REGION Network 2: Dose_Control_Linie_1
   IF "GDB_PLC".Start_Modus_Linie_1 AND NOT "GDB_PLC".Stop_Modus_Linie_1 THEN
       "FB_Dose_Control_DB_1"(Trigger_Start := "GDB_PLC".Dosierung_Start_Linie_1,   // "FB_Dose_Control"
                              Flow_Raw := "Tank 2 (Flow Meter)",
                              Target_Volume := "GDB_Getränk".Getränk_Linie_1.Dosiervolumen,
                              Not_Aus := "GDB_PLC".Not_Aus_Modus,
                              Discharge_Valve => "Tank 2 (Discharge Valve)",
                              Dosing_Status => "GDB_PLC".Dosing_Activate_Linie_1,
                              Füllmenge => "GDB_HMI".Füllmenge_Linie_1);
   END_IF;
END_REGION
END_ORGANIZATION_BLOCK

(* ===== HMI "HMI_RT_1" =====
system functions are stored by id; their names below are inferred from use
connection "HMI_Verbindung_1": ETHERNET, SMART_S7_1200_OMS

HMI tags "Standard-Variablentabelle"
   "Variable_Bildnummer" : UInt, internal
   "Start Button 1" : Bool = PLC "Start Button 1" AT %I5.0, 100 ms
   "Start Button 1 (Light)" : Bool = PLC "Start Button 1 (Light)" AT %Q4.4, 100 ms
   "Stop Button 1" : Bool = PLC "Stop Button 1" AT %I5.2, 100 ms
   "Emergency Stop 1" : Bool = PLC "Emergency Stop 1" AT %I3.7, 100 ms
   "GDB_PLC_Start_Modus" : Bool = PLC GDB_PLC.Start_Modus_Hauptleitung, 100 ms
   "GDB_PLC_Not_Aus_Modus" : Bool = PLC GDB_PLC.Not_Aus_Modus, 100 ms
   "GDB_HMI_Füllmenge" : Real = PLC GDB_HMI.Füllmenge_Linie_0, 100 ms
   "GDB_PLC_Dosing_Activate" : Bool = PLC GDB_PLC.Dosing_Activate_Linie_0, 100 ms
   "GDB_PLC_Füllventil_Stand" : Bool = PLC GDB_PLC.Füllventil_closed_Linie_0, 100 ms
   "Stop Button 1 (Light)" : Bool = PLC "Stop Button 1 (Light)" AT %Q4.6, 100 ms
   "GDB_HMI_Reset_Gesamtteile_0" : Bool = PLC GDB_HMI.Reset_Gesamtteile_0, 100 ms
   "GDB_HMI_Reset_Ausschluss_0" : Bool = PLC GDB_HMI.Reset_Ausschluss_0, 100 ms
   "GDB_PLC_Gesamtteile_Linie_0" : Int = PLC GDB_PLC.Gesamtteile_Linie_0, 100 ms
   "GDB_PLC_Altuell_Gewicht_Linie_0" : Real = PLC GDB_PLC.Altuell_Gewicht_Linie_0, 100 ms
   "GDB_PLC_Tankfüllvolumen" : Real = PLC GDB_PLC.Tankfüllvolumen_0, 100 ms
   "GDB_PLC_Dosiervolumen" : Real = PLC GDB_PLC.Dosiervolumen_0, 100 ms
   "GDB_Getränk_Getränk_Linie_1_VAR_Rezeptur_Datensatz" : Int = PLC GDB_Getränk.Getränk_Linie_1.VAR_Rezeptur_Datensatz, 100 ms
   "GDB_Getränk_Getränk_Linie_0_VAR_Rezeptur_Datensatz" : Int = PLC GDB_Getränk.Getränk_Linie_0.VAR_Rezeptur_Datensatz, 100 ms
   "GDB_Getränk_Getränk_Linie_0_VAR_Rezeptur" : Int = PLC GDB_Getränk.Getränk_Linie_0.VAR_Rezeptur, 100 ms
   "GDB_Getränk_Getränk_Linie_0_Tankfüllvolumen" : Real = PLC GDB_Getränk.Getränk_Linie_0.Tankfüllvolumen, 100 ms
   "GDB_Getränk_Getränk_Linie_0_Dosiervolumen" : Real = PLC GDB_Getränk.Getränk_Linie_0.Dosiervolumen, 100 ms
   "GDB_PLC_Tank_1_Level_norm" : Real = PLC GDB_PLC.Tank_1_Level_norm, 100 ms
   "Start Button 0" : Bool = PLC "Start Button 0" AT %I5.3, 100 ms
   "Stop Button 0" : Bool = PLC "Stop Button 0" AT %I5.1, 100 ms
   "Emergency Stop 0" : Bool = PLC "Emergency Stop 0" AT %I3.6, 100 ms
   "GDB_Getränk_Getränk_Linie_1_Tankfüllvolumen" : Real = PLC GDB_Getränk.Getränk_Linie_1.Tankfüllvolumen, 100 ms
   "GDB_Getränk_Getränk_Linie_1_Dosiervolumen" : Real = PLC GDB_Getränk.Getränk_Linie_1.Dosiervolumen, 100 ms
   "GDB_PLC_Tank_0_Level_norm" : Real = PLC GDB_PLC.Tank_0_Level_norm, 100 ms
   "GDB_PLC_Tankfüllvolumen_1" : Real = PLC GDB_PLC.Tankfüllvolumen_1, 100 ms
   "GDB_PLC_Dosiervolumen_1" : Real = PLC GDB_PLC.Dosiervolumen_1, 100 ms
   "GDB_PLC_Start_Modus_Linie_1" : Bool = PLC GDB_PLC.Start_Modus_Linie_1, 100 ms
   "GDB_PLC_Start_Modus_Linie_0" : Bool = PLC GDB_PLC.Start_Modus_Linie_0, 100 ms
   "GDB_PLC_Stop_Modus" : Bool = PLC GDB_PLC.Stop_Modus_Hauptleitung, 100 ms
   "GDB_HMI_NotAus_HMI" : Bool = PLC GDB_HMI.NotAus_HMI, 100 ms
   "Start Button 0 (Light)" : Bool = PLC "Start Button 0 (Light)" AT %Q4.3, 100 ms
   "GDB_PLC_Stop_Modus_Linie_0" : Bool = PLC GDB_PLC.Stop_Modus_Linie_0, 100 ms
   "GDB_PLC_Stop_Modus_Linie_1" : Bool = PLC GDB_PLC.Stop_Modus_Linie_1, 100 ms
   "GDB_PLC_Dosing_Activate_Linie_1" : Bool = PLC GDB_PLC.Dosing_Activate_Linie_1, 100 ms
   "GDB_HMI_Füllmenge_Linie_1" : Real = PLC GDB_HMI.Füllmenge_Linie_1, 100 ms
   "GDB_PLC_Altuell_Gewicht_Linie_1" : Real = PLC GDB_PLC.Altuell_Gewicht_Linie_1, 100 ms
   "GDB_PLC_Gesamtteile_Linie_1" : Int = PLC GDB_PLC.Gesamtteile_Linie_1, 100 ms
   "GDB_HMI_Reset_Gesamtteile_1" : Bool = PLC GDB_HMI.Reset_Gesamtteile_1, 100 ms
   "GDB_HMI_Reset_Ausschluss_1" : Bool = PLC GDB_HMI.Reset_Ausschluss_1, 100 ms
   "Benutzername" : WString[254], internal
   "GDB_Getränk_Getränk_Linie_1_VAR_Rezeptur" : Int = PLC GDB_Getränk.Getränk_Linie_1.VAR_Rezeptur, 100 ms
   "GDB_PLC_Ausschuss_Linie_1" : Int = PLC GDB_PLC.Ausschuss_Linie_1, 100 ms
   "GDB_PLC_Ausschuss_Linie_0" : Int = PLC GDB_PLC.Ausschuss_Linie_0, 100 ms
   "GDB_PLC_Anzahl_Paletten" : Int = PLC GDB_PLC.Anzahl_Paletten, 100 ms
   "GDB_PLC_Anzahl_Kanister_Packungbereich" : Int = PLC GDB_PLC.Anzahl_Kanister_Packungbereich, 100 ms
   "GDB_PLC_Anzahl_Kanister_Tr_Band_Halle_2" : Int = PLC GDB_PLC.Anzahl_Kanister_Tr_Band_Halle_2, 100 ms
   "GDB_PLC_Run_Hours" : Int = PLC GDB_PLC.Run_Hours, 100 ms
   "GDB_PLC_Run_Minutes" : Int = PLC GDB_PLC.Run_Minutes, 100 ms
   "GDB_PLC_Run_Seconds" : Int = PLC GDB_PLC.Run_Seconds, 100 ms
   "GDB_HMI_Meldung_Störung_HMI" : Int = PLC GDB_HMI.Meldung_HMI, 100 ms
   "GDB_HMI_Quittierung_Störung_HMI" : Int = PLC GDB_HMI.Quittierung_HMI, 100 ms
   "Störung_0" : Bool = PLC GDB_PLC.Störung[0] AT %DB1.DBX0.0, 100 ms
   "Störung_1" : Bool = PLC GDB_PLC.Störung[1] AT %DB1.DBX0.0, 100 ms
   "Störung_2" : Bool = PLC GDB_PLC.Störung[2] AT %DB1.DBX0.0, 100 ms
   "Störung_3" : Bool = PLC GDB_PLC.Störung[3] AT %DB1.DBX0.0, 100 ms
   "Störung_4" : Bool = PLC GDB_PLC.Störung[4] AT %DB1.DBX0.0, 100 ms
   "Störung_5" : Bool = PLC GDB_PLC.Störung[5] AT %DB1.DBX0.0, 100 ms
   "Störung_6" : Bool = PLC GDB_PLC.Störung[6] AT %DB1.DBX0.0, 100 ms
   "Störung_7" : Bool = PLC GDB_PLC.Störung[7] AT %DB1.DBX0.0, 100 ms
   "Störung_8" : Bool = PLC GDB_PLC.Störung[8] AT %DB1.DBX0.0, 100 ms
   "Störung_9" : Bool = PLC GDB_PLC.Störung[9] AT %DB1.DBX0.0, 100 ms
   "Störung_10" : Bool = PLC GDB_PLC.Störung[10] AT %DB1.DBX0.0, 100 ms
   "Störung_15" : Bool = PLC GDB_PLC.Störung[15] AT %DB1.DBX0.0, 100 ms
   "Störung_14" : Bool = PLC GDB_PLC.Störung[14] AT %DB1.DBX0.0, 100 ms
   "Störung_13" : Bool = PLC GDB_PLC.Störung[13] AT %DB1.DBX0.0, 100 ms
   "Störung_12" : Bool = PLC GDB_PLC.Störung[12] AT %DB1.DBX0.0, 100 ms
   "Störung_16" : Bool = PLC GDB_PLC.Störung[16] AT %DB1.DBX0.0, 100 ms
   "Störung_11" : Bool = PLC GDB_PLC.Störung[11] AT %DB1.DBX0.0, 100 ms
   "Haupt_Stop_HMI" : Bool = PLC GDB_HMI.Haupt_Stop_HMI AT %DB1.DBX0.0, 100 ms

discrete alarms
   1: 'Störung_AbfüllLinie_0_Tr_Band_0', class Störung, trigger "GDB_HMI_Meldung_Störung_HMI" bit 0
   2: 'Störung_AbfüllMaschine_0', class Störung, trigger "GDB_HMI_Quittierung_Störung_HMI" bit 1
   3: 'Störung_AbfüllMaschine_1', class Störung, trigger "GDB_HMI_Quittierung_Störung_HMI" bit 2
   4: 'Störung_Gewichtkontrolle_Linie_0', class Störung, trigger "GDB_HMI_Quittierung_Störung_HMI" bit 3
   5: 'Störung_Gewichtkontrolle_Linie_1', class Störung, trigger "GDB_HMI_Quittierung_Störung_HMI" bit 4
   6: 'Störung_Hauptlinie_Kurvenband_0', class Störung, trigger "GDB_HMI_Meldung_Störung_HMI" bit 5
   7: 'Störung_Hauptlinie_Band_1', class Störung, trigger "GDB_HMI_Meldung_Störung_HMI" bit 6
   8: 'Störung_Hauptlinie_Band_2', class Störung, trigger "GDB_HMI_Meldung_Störung_HMI" bit 7
   9: 'Störung_Hauptlinie_T - Band_3', class Störung, trigger "GDB_HMI_Meldung_Störung_HMI" bit 8
   10: 'Störung_Hauptlinie_Band_4', class Störung, trigger "GDB_HMI_Meldung_Störung_HMI" bit 9
   11: 'Störung_Hauptlinie_Kurvenband_1', class Störung, trigger "GDB_HMI_Meldung_Störung_HMI" bit 10
   12: 'Störung_Sortierabschnitt', class Störung, trigger "GDB_HMI_Meldung_Störung_HMI" bit 11
   13: 'Störung_Transport_Band_1_PackungLinie_0', class Störung, trigger "GDB_HMI_Meldung_Störung_HMI" bit 12
   14: 'Störung_Transport_Band_2_PackungLinie_0', class Störung, trigger "GDB_HMI_Meldung_Störung_HMI" bit 13
   15: 'Störung_Band mit Positionierleisten', class Störung, trigger "GDB_HMI_Meldung_Störung_HMI" bit 14
   17: 'Störung_Pick & Place_Linie_0', class Störung, trigger "GDB_HMI_Meldung_Störung_HMI" bit 15

text list "Rezepturen_Linie_0": 2 'Gurkenlimonade, 7L'; 4 'Gurkenlimonade, 5L'

text list "Rezepturen_Linie_1": 1 'Lavendel-Limonade, 5L'; 2 'Lavendel-Limonade, 8L'

recipe "Linie_0": Tankfüllvolumen <- "GDB_Getränk_Getränk_Linie_0_Tankfüllvolumen", Dosiervolumen <- "GDB_Getränk_Getränk_Linie_0_Dosiervolumen"

recipe "Linie_1": Tankfüllvolumen <- "GDB_Getränk_Getränk_Linie_1_Tankfüllvolumen", Dosiervolumen <- "GDB_Getränk_Getränk_Linie_1_Dosiervolumen"

Template "Vorlage_1" 800x480
   Button "Exit" at 722,440 size 55x39; TextOff 'Exit'; PictureOff "ExitRuntime_KTP900_Basic_PN_TR"; PictureOn "ExitRuntime_KTP900_Basic_PN_TR"
      on Release: StopRuntime(0)
   Button "Log on" at 622,440 size 55x39; TextOff 'Log on'; PictureOff "Login_KTP900_Basic_PN_TR"; PictureOn "Login_KTP900_Basic_PN_TR"
      on Press: ActivateScreen("Benutzerverwaltung", 0)
   Button "Template_Button" at 522,440 size 55x39; TextOff 'Rezept'; PictureOff "Rezeptur_mono"
      on Press: ActivateScreen("Rezepturen", 0)
   Button "Template_Button_1" at 422,440 size 55x39; TextOff 'Putz'
      on Click: function_be740847(30)
   Button "Template_Button_2" at 322,440 size 55x39; TextOff 'Text'; PictureOff "Navigates to Systembilder for KTP900 Basic+ PN 17.0.0.0"
      on Click: ActivateScreen("Systembilder", 0)
   Button "Template_Button_3" at 222,440 size 55x39; TextOff 'Übers'; PictureOff "Navigates to Systembilder for KTP900 Basic+ PN 17.0.0.0"
      on Press: ActivateScreen("Übersicht", 0)
   Button "Start screen" at 122,440 size 55x39; TextOff 'Abfüll'; TextOn 'Start screen'; PictureOff "NavigateHome_KTP900_Basic_PN_TR"; PictureOn "NavigateHome_KTP900_Basic_PN_TR"
      on Press: ActivateScreen("Abfüllbereich", 0)
   Button "Alarms" at 22,440 size 55x39; TextOff 'Alarms'; PictureOff "AlarmDisplay_KTP900_Basic_PN_TR"; PictureOn "AlarmDisplay_KTP900_Basic_PN_TR"
      on Press: ActivateScreen("Meldungen", 0)
   SymbolicIOField "Symbolisches_EA_Feld_Bild" at 73,7 size 620x26; TextOff '0'; TextOn '1'; TextList "TextList_ScreenNames"
      ProcessValue <- "Variable_Bildnummer"
      on Change: ActivateScreenByNumber("Variable_Bildnummer", 0)
   DateTimeField "HmiScreenItemData" at 695,20 size 105x20
   DateTimeField "HmiScreenItemData_1" at 695,0 size 105x20
   GraphicView "Logo" at 0,0 size 71x40; Picture "Logo of HMI_1"
   GraphicView "Vorlage_Grafikanzeige_1" at 425,42 size 23x23; Picture "login-icon-3060"
   IOField "Vorlage_EA-Feld_1" at 489,44 size 90x19; FormatPattern ????????????????????????????????????????????????????????????????????????????????
      ProcessValue <- "Benutzername"
   Button "Schaltfläche_1" at 590,44 size 90x19; TextOff 'Anmelden'
      on Press: function_a2a04561()
   Button "Schaltfläche_2" at 697,44 size 90x19; TextOff 'Abmelden'
      on Press: function_f23ef4c9()

screen "Abfüllbereich" 800x480, template "Vorlage_1"
   on GenerateScreen: SetTag("Variable_Bildnummer", 1)
   GraphicView "Grafikanzeige_3" at 461,260 size 29x32; Picture "Ventil_Green-removebg-preview"
   GraphicView "Grafikanzeige_4" at 461,260 size 29x32; Picture "Ventil_Gray-removebg-preview"
      Visibility <- "GDB_PLC_Dosing_Activate"
   Bar "Balken_3" at 454,338 size 34x40; MinimumValue 0; MaximumValue 10
      ProcessValue <- "GDB_HMI_Füllmenge"
   GraphicView "Grafikanzeige_6" at 452,317 size 38x63; Picture "Bottle_1"
   Button "Schaltfläche_7" at 707,356 size 72x26; TextOff 'Reset'
      Appearance <- "GDB_HMI_Reset_Gesamtteile_0"
      on Press: SetBit("GDB_HMI_Reset_Gesamtteile_0")
      on Release: ResetBit("GDB_HMI_Reset_Gesamtteile_0")
   Button "Schaltfläche_5" at 708,395 size 72x28; TextOff 'Reset'
      Appearance <- "GDB_HMI_Reset_Ausschluss_0"
      on Press: SetBit("GDB_HMI_Reset_Ausschluss_0")
      on Release: ResetBit("GDB_HMI_Reset_Ausschluss_0")
   TextField "Textfeld_20" at 639,147 size 113x17; Text 'Die Linie ist in Betrieb,'
   TextField "Textfeld_21" at 612,158 size 175x17; Text 'ein Rezeptwechsel ist nicht möglich'
   GraphicView "Grafikanzeige_7" at 323,260 size 29x32; Picture "Ventil_Green-removebg-preview"
   GraphicView "Grafikanzeige_8" at 323,260 size 29x32; Picture "Ventil_Gray-removebg-preview"
      Visibility <- "GDB_PLC_Dosing_Activate_Linie_1"
   Button "Schaltfläche_10" at 179,356 size 72x26; TextOff 'Reset'
      on Release: ResetBit("GDB_HMI_Reset_Gesamtteile_1")
      on Press: SetBit("GDB_HMI_Reset_Gesamtteile_1")
      Appearance <- "GDB_HMI_Reset_Gesamtteile_0"
   Button "Schaltfläche_11" at 180,395 size 72x28; TextOff 'Reset'
      on Release: ResetBit("GDB_HMI_Reset_Ausschluss_1")
      on Press: SetBit("GDB_HMI_Reset_Ausschluss_1")
      Appearance <- "GDB_HMI_Reset_Ausschluss_0"
   TextField "Textfeld_41" at 41,146 size 113x17; Text 'Die Linie ist in Betrieb,'
   TextField "Textfeld_42" at 14,157 size 175x17; Text 'ein Rezeptwechsel ist nicht möglich'
   Bar "Balken_6" at 318,338 size 34x40; MinimumValue 0; MaximumValue 10
      ProcessValue <- "GDB_HMI_Füllmenge_Linie_1"
   GraphicView "Grafikanzeige_10" at 316,317 size 38x63; Picture "Bottle_1"
   TextField "Textfeld_22" at 138,69 size 162x20; Text 'ABFÜLLMASCHINE Linie 1'
   Button "Schaltfläche_6" at 201,111 size 89x32; TextOff 'Start'; Authorization "Bedienen"
      on Press: SetBit("Start Button 1")
      Appearance <- "Start Button 1 (Light)"
   Button "Schaltfläche_8" at 296,111 size 89x32; TextOff 'Stop'
      on Click: ResetBit("Stop Button 1")
      Appearance <- "GDB_PLC_Stop_Modus_Linie_1"
   TextField "Textfeld_1" at 538,69 size 162x20; Text 'ABFÜLLMASCHINE Linie 0'
   Button "Schaltfläche_1" at 511,111 size 89x32; TextOff 'Start'; Authorization "Bedienen"
      on Press: SetBit("Start Button 0")
      Appearance <- "Start Button 0 (Light)"
   Button "Schaltfläche_2" at 414,111 size 89x32; TextOff 'Stop'
      on Click: ResetBit("Stop Button 0")
      Appearance <- "GDB_PLC_Stop_Modus_Linie_0"
   Button "Schaltfläche_3" at 290,403 size 225x34; TextOff 'NOT AUS'
      Appearance <- "GDB_PLC_Not_Aus_Modus"
      on Press: InvertBit("GDB_HMI_NotAus_HMI")
   Bar "Balken_2" at 437,171 size 37x62; MinimumValue 0; MaximumValue 300
      ProcessValue <- "GDB_PLC_Tank_0_Level_norm"
   GraphicView "Grafikanzeige_5" at 460,247 size 25x19; Picture "Grafik_6"
   Rectangle "Rechteck_2" at 468,292 size 6x44
      Visibility <- "GDB_PLC_Dosing_Activate"
   Group "Group" at 461,260 size 29x32; Picture "Ventil_Green-removebg-preview"
   GraphicView "Grafikanzeige_2" at 427,154 size 89x101; Picture "rzhbt5dt.1cr"
   Group "Group_3" at 452,317 size 38x63; Picture "Bottle_1"
   SymbolicIOField "Symbolisches EA-Feld_1" at 615,121 size 164x20; TextOff '0'; TextOn '1'; TextList "Rezepturen_Linie_0"
      ProcessValue <- "GDB_Getränk_Getränk_Linie_0_VAR_Rezeptur_Datensatz"
   TextField "Textfeld_2" at 670,101 size 51x20; Text 'Rezept'
   Group "Group_4" at 612,147 size 175x28
   Button "Schaltfläche_4" at 610,150 size 175x23; TextOff 'Rezept hochladen'; Authorization "Bedienen"
      on Click: function_eba64363("Linie_0", "GDB_Getränk_Getränk_Linie_0_VAR_Rezeptur_Datensatz", 1, N)
      Visibility <- "GDB_PLC_Start_Modus_Linie_0"
   TextField "Textfeld_3" at 543,260 size 70x22; Text 'Füllmenge'
   TextField "Textfeld_19" at 765,293 size 19x20; Text 'Kg'
   TextField "Textfeld_4" at 550,230 size 61x22; Text 'Füllstand'
   TextField "Textfeld_7" at 676,233 size 11x20; Text 'L'
   TextField "Textfeld_12" at 643,185 size 44x20; Text 'Daten'
   IOField "EA-Feld_4" at 708,229 size 59x26; FormatPattern 999
      ProcessValue <- "GDB_PLC_Tank_0_Level_norm"
   TextField "Textfeld_10" at 555,291 size 55x22; Text 'Gewicht'
   TextField "Textfeld_11" at 712,205 size 51x22; Text 'Istwert'
   TextField "Textfeld_15" at 619,206 size 53x22; Text 'Sollwert'
   IOField "EA-Feld_7" at 708,261 size 59x26; FormatPattern 9.9
      ProcessValue <- "GDB_HMI_Füllmenge"
   IOField "EA-Feld_8" at 708,291 size 59x26; FormatPattern 9.9
      ProcessValue <- "GDB_PLC_Altuell_Gewicht_Linie_0"
   TextField "Textfeld_8" at 677,262 size 11x20; Text 'L'
   TextField "Textfeld_16" at 767,233 size 11x20; Text 'L'
   TextField "Textfeld_17" at 766,264 size 11x20; Text 'L'
   TextField "Textfeld_18" at 676,293 size 19x20; Text 'Kg'
   IOField "EA-Feld_9" at 619,229 size 59x26; FormatPattern 999
      ProcessValue <- "GDB_PLC_Tankfüllvolumen"
   IOField "EA-Feld_10" at 619,260 size 59x26; FormatPattern 9.9
      ProcessValue <- "GDB_PLC_Dosiervolumen"
   IOField "EA-Feld_11" at 619,291 size 59x26; FormatPattern 9.9
      ProcessValue <- "GDB_PLC_Dosiervolumen"
   Bar "Balken_5" at 301,179 size 37x52; MinimumValue 0; MaximumValue 300
      ProcessValue <- "GDB_PLC_Tank_1_Level_norm"
   GraphicView "Grafikanzeige_1" at 322,248 size 25x19; Picture "Grafik_6"
   GraphicView "Grafikanzeige_9" at 290,156 size 89x101; Picture "rzhbt5dt.1cr"
   Rectangle "Rechteck_11" at 332,292 size 6x44
      Visibility <- "GDB_PLC_Dosing_Activate_Linie_1"
   Group "Group_9" at 323,260 size 29x32; Picture "Ventil_Green-removebg-preview"
   Group "Group_16" at 316,317 size 38x63; Picture "Bottle_1"
   SymbolicIOField "Symbolisches EA-Feld_2" at 17,121 size 164x20; TextOn '1'; TextOff '0'; TextList "Rezepturen_Linie_1"
      ProcessValue <- "GDB_Getränk_Getränk_Linie_1_VAR_Rezeptur_Datensatz"
   TextField "Textfeld_40" at 72,101 size 51x20; Text 'Rezept'
   Group "Group_14" at 14,146 size 175x28
   Button "Schaltfläche_12" at 12,150 size 175x23; TextOff 'Rezept hochladen'; Authorization "Bedienen"
      on Click: function_eba64363("Linie_1", "GDB_Getränk_Getränk_Linie_1_VAR_Rezeptur_Datensatz", 1, N)
      Visibility <- "GDB_PLC_Start_Modus_Linie_1"
   TextField "Textfeld_28" at 15,259 size 70x22; Text 'Füllmenge'
   TextField "Textfeld_29" at 237,293 size 19x20; Text 'Kg'
   TextField "Textfeld_30" at 22,230 size 61x22; Text 'Füllstand'
   TextField "Textfeld_31" at 148,233 size 11x20; Text 'L'
   TextField "Textfeld_32" at 115,185 size 44x20; Text 'Daten'
   IOField "EA-Feld_6" at 180,229 size 59x26; FormatPattern 999
      ProcessValue <- "GDB_PLC_Tank_1_Level_norm"
   TextField "Textfeld_33" at 27,291 size 55x22; Text 'Gewicht'
   TextField "Textfeld_34" at 184,205 size 51x22; Text 'Istwert'
   TextField "Textfeld_35" at 91,206 size 53x22; Text 'Sollwert'
   IOField "EA-Feld_12" at 180,260 size 59x26; FormatPattern 9.9
      ProcessValue <- "GDB_HMI_Füllmenge_Linie_1"
   IOField "EA-Feld_13" at 180,291 size 59x26; FormatPattern 9.9
      ProcessValue <- "GDB_PLC_Altuell_Gewicht_Linie_1"
   TextField "Textfeld_36" at 149,262 size 11x20; Text 'L'
   TextField "Textfeld_37" at 239,233 size 11x20; Text 'L'
   TextField "Textfeld_38" at 238,264 size 11x20; Text 'L'
   TextField "Textfeld_39" at 148,292 size 19x20; Text 'Kg'
   IOField "EA-Feld_14" at 91,229 size 59x26; FormatPattern 999
      ProcessValue <- "GDB_PLC_Tankfüllvolumen_1"
   IOField "EA-Feld_15" at 91,260 size 59x26; FormatPattern 9.9
      ProcessValue <- "GDB_PLC_Dosiervolumen_1"
   IOField "EA-Feld_16" at 91,290 size 59x26; FormatPattern 9.9
      ProcessValue <- "GDB_PLC_Dosiervolumen_1"
   TextField "Textfeld_23" at 20,360 size 56x22; Text 'Gesamt'
   TextField "Textfeld_24" at 21,400 size 73x22; Text 'Ausschuss'
   IOField "EA-Feld_1" at 100,359 size 47x26; FormatPattern 999
      ProcessValue <- "GDB_PLC_Gesamtteile_Linie_1"
   TextField "Textfeld_25" at 75,328 size 113x20; Text 'Produktiondaten'
   IOField "EA-Feld_2" at 101,400 size 47x26; FormatPattern 9999
      ProcessValue <- "GDB_PLC_Ausschuss_Linie_1"
   TextField "Textfeld_26" at 146,362 size 30x20; Text 'Kan.'
   TextField "Textfeld_27" at 147,403 size 30x20; Text 'Kan.'
   Group "Group_10" at 179,356 size 74x30
   Group "Group_11" at 180,395 size 74x32
   TextField "Textfeld_5" at 549,360 size 56x22; Text 'Gesamt'
   TextField "Textfeld_6" at 549,400 size 73x22; Text 'Ausschuss'
   IOField "EA-Feld_3" at 628,359 size 47x26; FormatPattern 9999
      ProcessValue <- "GDB_PLC_Gesamtteile_Linie_0"
   TextField "Textfeld_9" at 603,328 size 113x20; Text 'Produktiondaten'
   IOField "EA-Feld_5" at 629,400 size 47x26; FormatPattern 9999
      ProcessValue <- "GDB_PLC_Ausschuss_Linie_0"
   TextField "Textfeld_13" at 674,362 size 30x20; Text 'Kan.'
   TextField "Textfeld_14" at 675,403 size 30x20; Text 'Kan.'
   Group "Group_2" at 707,356 size 74x30
   Group "Group_1" at 708,395 size 74x32

screen "Systembilder" 800x480, template "Vorlage_1"
   on GenerateScreen: SetTag("Variable_Bildnummer", 2)
   Button "Back" at 1,41 size 159x47; TextOff 'Back'
      on Release: ActivateScreen("Abfüllbereich", 0)
   Button "HmiScreenItemData" at 36,195 size 159x47; TextOff 'SIMATIC PLC system diagnos...'; PictureOff "Navigates to SIMATIC PLC Systemdiagnose for KTP900 Basic+ PN 17.0.0.0"; PictureOn "Navigates to SIMATIC PLC Systemdiagnose for KTP900 Basic+ PN 17.0.0.0"
      on Release: ActivateScreen("SIMATIC PLC Systemdiagnose", 0)
   Button "HmiScreenItemData_2" at 36,253 size 159x47; TextOff 'User administration'; PictureOff "Navigates to Benutzerverwaltung for KTP900 Basic+ PN 17.0.0.0"; PictureOn "Navigates to Benutzerverwaltung for KTP900 Basic+ PN 17.0.0.0"
      on Release: ActivateScreen("Benutzerverwaltung", 0)
   Button "HmiScreenItemData_3" at 36,312 size 159x47; TextOff 'System information'; PictureOff "Navigates to Systeminformationen for KTP900 Basic+ PN 17.0.0.0"; PictureOn "Navigates to Systeminformationen for KTP900 Basic+ PN 17.0.0.0"
      on Release: ActivateScreen("Systeminformationen", 0)

screen "SIMATIC PLC Systemdiagnose" 800x480, template "Vorlage_1"
   on GenerateScreen: SetTag("Variable_Bildnummer", 3)
   SysDiagControl "HmiScreenItemData" at 1,89 size 796x343
   Button "Back" at 1,41 size 159x47; TextOff 'Back'
      on Release: ActivateScreen("Systembilder", 0)

screen "Projektinformationen" 800x480, template "Vorlage_1"
   on GenerateScreen: SetTag("Variable_Bildnummer", 4)
   TextField "HmiScreenItemData" at 35,91 size 171x28; Text 'Project name:'
   TextField "HmiScreenItemData_1" at 241,91 size 524x28; Text 'Projekt_10'
   TextField "HmiScreenItemData_2" at 35,121 size 171x28; Text 'Created on:'
   TextField "HmiScreenItemData_3" at 241,121 size 524x28; Text '07.04.2016 11:51:36'
   TextField "HmiScreenItemData_4" at 35,151 size 171x28; Text 'Author:'
   TextField "HmiScreenItemData_5" at 241,151 size 524x28; Text 'Matthias Habermann'
   TextField "HmiScreenItemData_6" at 35,181 size 171x28; Text 'Description:'
   TextField "HmiScreenItemData_7" at 241,181 size 524x28; Text '(not configured)'
   Button "Back" at 1,41 size 159x47; TextOff 'Back'
      on Release: ActivateScreen("Systembilder", 0)

screen "Benutzerverwaltung" 800x480, template "Vorlage_1"
   on GenerateScreen: SetTag("Variable_Bildnummer", 5)
   UserView "HmiScreenItemData" at 1,89 size 796x343
   Button "Back" at 1,41 size 159x47; TextOff 'Back'
      on Release: ActivateScreen("Systembilder", 0)

screen "Systeminformationen" 800x480, template "Vorlage_1"
   on GenerateScreen: SetTag("Variable_Bildnummer", 6)
   TextField "HmiScreenItemData" at 35,91 size 171x28; Text 'HMI device type:'
   TextField "HmiScreenItemData_1" at 241,91 size 524x28; Text 'KTP900 Basic+ PN 17.0.0.0'
   TextField "HmiScreenItemData_2" at 35,121 size 171x28; Text 'Connection:'
   TextField "HmiScreenItemData_3" at 241,121 size 524x28; Text 'PROFINET (X1)'
   TextField "HmiScreenItemData_4" at 35,151 size 171x28; Text 'PLC:'
   TextField "HmiScreenItemData_5" at 241,151 size 524x28; Text 'SIMATIC S7 1200'
   Button "Back" at 1,41 size 159x47; TextOff 'Back'
      on Release: ActivateScreen("Systembilder", 0)

screen "Rezepturen" 800x480, template "Vorlage_1"
   on GenerateScreen: SetTag("Variable_Bildnummer", 8)
   RecipeView "Rezepturanzeige_1" at 24,111 size 376x322; DataRecordNameCaption 'Dosiervolumen'; Tag4DataRecord "GDB_Getränk_Getränk_Linie_0_VAR_Rezeptur_Datensatz"; Tag4RecipeNumber "GDB_Getränk_Getränk_Linie_0_VAR_Rezeptur"; Recipe "Linie_0"
   Button "Back" at 24,47 size 159x47; TextOn 'Back'; TextOff 'Back'
      on Release: ActivateScreen("Abfüllbereich", 0)
   RecipeView "Rezepturanzeige_2" at 406,111 size 376x322; DataRecordNameCaption 'Dosiervolumen'; Recipe "Linie_1"; Tag4RecipeNumber "GDB_Getränk_Getränk_Linie_1_VAR_Rezeptur"; Tag4DataRecord "GDB_Getränk_Getränk_Linie_1_VAR_Rezeptur_Datensatz"

screen "Verschiedene Aufgaben" 800x480, template "Vorlage_1"
   on GenerateScreen: SetTag("Variable_Bildnummer", 7)
   Button "Online" at 36,135 size 159x47; TextOff 'Online'
      on Release: function_bb44b551(0)
   Button "Offline" at 36,194 size 159x47; TextOff 'Offline'
      on Release: function_bb44b551(1)
   Button "Transfer" at 36,253 size 159x47; TextOff 'Transfer'
      on Release: function_bb44b551(2)
   Button "Toggle language" at 36,312 size 159x47; TextOff 'Toggle language'
      on Release: function_fb9197e8(-1)
   Button "Stop Runtime" at 36,371 size 159x47; TextOff 'Stop Runtime'
      on Release: StopRuntime(0)
   Button "Back" at 1,41 size 159x47; TextOff 'Back'
      on Release: ActivateScreen("Systembilder", 0)

screen "Meldungen" 800x480, template "Vorlage_1"
   on GenerateScreen: SetTag("Variable_Bildnummer", 9)
   AlarmView "Meldeanzeige_1" at 11,71 size 781x322
   Button "Schaltfläche_1" at 573,400 size 143x26; TextOff 'Meldungen löschen'
      on Click: function_e14cd482(0)

screen "Übersicht" 800x480, template "Vorlage_1"
   on GenerateScreen: SetTag("Variable_Bildnummer", 10)
   IOField "EA-Feld_4" at 166,174 size 59x26; FormatPattern 999
      ProcessValue <- "GDB_PLC_Tank_0_Level_norm"
   IOField "EA-Feld_3" at 166,202 size 59x26; FormatPattern 999
      ProcessValue <- "GDB_PLC_Gesamtteile_Linie_0"
   IOField "EA-Feld_5" at 166,230 size 59x26; FormatPattern 999
      ProcessValue <- "GDB_PLC_Ausschuss_Linie_0"
   Group "Group_4" at 178,152 size 77x18
   TextField "Textfeld_46" at 17,152 size 114x20; Text 'Abfüllmaschine 0'
   TextField "Textfeld_47" at 17,176 size 89x22; Text 'Tanrfüllstand'
   TextField "Textfeld_48" at 17,201 size 56x22; Text 'Gesamt'
   TextField "Textfeld_49" at 17,228 size 73x22; Text 'Ausschuss'
   TextField "Textfeld_50" at 227,209 size 30x20; Text 'Kan.'
   TextField "Textfeld_51" at 227,236 size 30x20; Text 'Kan.'
   TextField "Textfeld_52" at 227,182 size 11x20; Text 'L'
   Circle "Kreis_3" at 178,155 size 12x12
      Visibility <- "GDB_PLC_Start_Modus_Linie_0"
   TextField "Textfeld_43" at 196,152 size 59x18; Text 'In Betrieb'
      Visibility <- "GDB_PLC_Start_Modus_Linie_0"
   Group "Group_5" at 178,152 size 77x18
   Group "Group_7" at 178,152 size 77x18
   Group "Group" at 178,152 size 77x18
   Circle "Kreis_5" at 178,155 size 12x12
      Visibility <- "GDB_PLC_Stop_Modus_Linie_0"
   TextField "Textfeld_44" at 199,152 size 56x18; Text 'Gestoppt'
      Visibility <- "GDB_PLC_Stop_Modus_Linie_0"
   TextField "Textfeld_45" at 198,152 size 57x18; Text 'NOT AUS'
      Visibility <- "GDB_PLC_Not_Aus_Modus"
   Circle "Kreis_6" at 178,155 size 12x12
      Visibility <- "GDB_PLC_Not_Aus_Modus"
   Circle "Kreis_7" at 711,156 size 12x12
      Visibility <- "GDB_PLC_Stop_Modus_Linie_1"
   TextField "Textfeld_4" at 732,153 size 56x18; Text 'Gestoppt'
      Visibility <- "GDB_PLC_Stop_Modus_Linie_1"
   TextField "Textfeld_5" at 730,153 size 57x18; Text 'NOT AUS'
      Visibility <- "GDB_PLC_Not_Aus_Modus"
   Circle "Kreis_8" at 710,156 size 12x12
      Visibility <- "GDB_PLC_Not_Aus_Modus"
   Group "Group_9" at 710,153 size 77x18
   Group "Group_10" at 710,153 size 77x18
   Group "Group_6" at 711,153 size 77x18
   Circle "Kreis_9" at 710,156 size 12x12
      Visibility <- "GDB_PLC_Start_Modus_Linie_1"
   TextField "Textfeld_6" at 728,153 size 59x18; Text 'In Betrieb'
      Visibility <- "GDB_PLC_Start_Modus_Linie_1"
   TextField "Textfeld_17" at 199,271 size 57x18; Text 'NOT AUS'
      Visibility <- "GDB_PLC_Not_Aus_Modus"
   Circle "Kreis_12" at 179,274 size 12x12
      Visibility <- "GDB_PLC_Not_Aus_Modus"
   Group "Group_16" at 179,271 size 77x18
   Group "Group_20" at 179,271 size 77x18
   Group "Group_19" at 179,271 size 77x18
   Circle "Kreis_13" at 179,274 size 12x12
      Visibility <- "GDB_PLC_Start_Modus_Linie_1"
   TextField "Textfeld_18" at 197,271 size 59x18; Text 'In Betrieb'
      Visibility <- "GDB_PLC_Start_Modus_Linie_1"
   Group "Group_17" at 179,271 size 77x18
   Group "Group_18" at 179,271 size 77x18
   Circle "Kreis_15" at 179,274 size 12x12
      Visibility <- "GDB_PLC_Stop_Modus"
   TextField "Textfeld_24" at 200,271 size 56x18; Text 'Gestoppt'
      Visibility <- "GDB_PLC_Stop_Modus"
   TextField "Textfeld_22" at 199,271 size 57x18; Text 'NOT AUS'
      Visibility <- "GDB_PLC_Not_Aus_Modus"
   Circle "Kreis_14" at 179,274 size 12x12
      Visibility <- "GDB_PLC_Not_Aus_Modus"
   Circle "Kreis_16" at 179,274 size 12x12
      Visibility <- "GDB_PLC_Start_Modus"
   TextField "Textfeld_25" at 197,271 size 59x18; Text 'In Betrieb'
      Visibility <- "GDB_PLC_Start_Modus"
   TextField "Textfeld_27" at 198,363 size 57x18; Text 'NOT AUS'
      Visibility <- "GDB_PLC_Not_Aus_Modus"
   Circle "Kreis_17" at 178,366 size 12x12
      Visibility <- "GDB_PLC_Not_Aus_Modus"
   Group "Group_22" at 178,363 size 77x18
   Group "Group_26" at 178,364 size 77x18
   Group "Group_25" at 178,363 size 77x18
   Circle "Kreis_18" at 178,366 size 12x12
      Visibility <- "GDB_PLC_Start_Modus_Linie_1"
   TextField "Textfeld_28" at 196,363 size 59x18; Text 'In Betrieb'
      Visibility <- "GDB_PLC_Start_Modus_Linie_1"
   Group "Group_23" at 178,363 size 77x18
   Group "Group_24" at 178,363 size 77x18
   Circle "Kreis_20" at 178,366 size 12x12
      Visibility <- "GDB_PLC_Stop_Modus"
   TextField "Textfeld_30" at 199,363 size 56x18; Text 'Gestoppt'
      Visibility <- "GDB_PLC_Stop_Modus"
   TextField "Textfeld_29" at 198,363 size 57x18; Text 'NOT AUS'
      Visibility <- "GDB_PLC_Not_Aus_Modus"
   Circle "Kreis_19" at 178,366 size 12x12
      Visibility <- "GDB_PLC_Not_Aus_Modus"
   Circle "Kreis_21" at 178,367 size 12x12
      Visibility <- "GDB_PLC_Start_Modus"
   TextField "Textfeld_31" at 196,364 size 59x18; Text 'In Betrieb'
      Visibility <- "GDB_PLC_Start_Modus"
   Group "Group_11" at 8,151 size 250x108
   IOField "EA-Feld_2" at 699,203 size 59x26; FormatPattern 999
      ProcessValue <- "GDB_PLC_Gesamtteile_Linie_1"
   IOField "EA-Feld_6" at 699,231 size 59x26; FormatPattern 999
      ProcessValue <- "GDB_PLC_Ausschuss_Linie_1"
   TextField "Textfeld_10" at 550,153 size 114x20; Text 'Abfüllmaschine 1'
   TextField "Textfeld_11" at 550,177 size 89x22; Text 'Tanrfüllstand'
   TextField "Textfeld_12" at 550,202 size 56x22; Text 'Gesamt'
   TextField "Textfeld_13" at 550,229 size 73x22; Text 'Ausschuss'
   TextField "Textfeld_14" at 760,210 size 30x20; Text 'Kan.'
   TextField "Textfeld_15" at 760,237 size 30x20; Text 'Kan.'
   TextField "Textfeld_16" at 760,183 size 11x20; Text 'L'
   IOField "EA-Feld_1" at 698,176 size 59x26; FormatPattern 999
      ProcessValue <- "GDB_PLC_Tank_1_Level_norm"
   IOField "EA-Feld_7" at 166,294 size 59x26; FormatPattern 999
      ProcessValue <- "GDB_PLC_Anzahl_Kanister_Packungbereich"
   IOField "EA-Feld_8" at 166,322 size 59x26; FormatPattern 999
      ProcessValue <- "GDB_PLC_Anzahl_Paletten"
   TextField "Textfeld_19" at 17,271 size 114x20; Text 'Packungsbereich'
   TextField "Textfeld_20" at 17,295 size 104x22; Text 'Anzahl Kanister'
   TextField "Textfeld_21" at 17,320 size 104x22; Text 'Anzahl Paletten'
   TextField "Textfeld_23" at 225,299 size 30x20; Text 'Kan.'
   TextField "Textfeld_9" at 225,327 size 26x20; Text 'Pal.'
   Group "Group_2" at 179,271 size 77x18
   TextField "Textfeld_26" at 16,363 size 145x20; Text 'Förderband zu Halle 2'
   TextField "Textfeld_32" at 16,386 size 104x22; Text 'Anzahl Kanister'
   IOField "EA-Feld_9" at 165,387 size 59x26; FormatPattern 999
      ProcessValue <- "GDB_PLC_Anzahl_Kanister_Tr_Band_Halle_2"
   TextField "Textfeld_33" at 222,392 size 30x20; Text 'Kan.'
   Group "Group_1" at 178,363 size 77x19
   Group "Group_3" at 710,153 size 78x18
   GraphicView "Grafikanzeige_1" at 264,147 size 279x279; Picture "Screenshot_2026-05-19_171715-removebg-preview"
   Group "Group_12" at 8,76 size 786x61
   Rectangle "Rechteck_7" at 7,76 size 786x61
      Visibility <- "GDB_PLC_Start_Modus"
   Group "Group_8" at 276,86 size 296x50
   Group "Group_13" at 7,76 size 786x61
   Group "Group_21" at 380,375 size 61x17
   Group "Group_28" at 509,333 size 63x17
   Group "Group_14" at 381,333 size 61x17
   Group "Group_15" at 380,295 size 61x17
   Group "Group_27" at 505,289 size 63x17
   TextField "Textfeld_41" at 448,242 size 50x17; Text 'Störung'
      Visibility <- "Störung_7"
   Ellipse "Ellipse_9" at 465,274 size 9x9
      Visibility <- "Störung_7"
   Group "Group_31" at 413,255 size 50x28
   TextField "Textfeld_53" at 476,255 size 50x17; Text 'Störung'
      Visibility <- "Störung_6"
   Ellipse "Ellipse_7" at 486,274 size 9x9
      Visibility <- "Störung_6"
   TextField "Textfeld_55" at 369,281 size 50x17; Text 'Störung'
      Visibility <- "Störung_9"
   Ellipse "Ellipse_10" at 396,273 size 9x9
      Visibility <- "Störung_9"
   Ellipse "Ellipse_6" at 375,254 size 9x9
      Visibility <- "Störung_15"
   TextField "Textfeld_42" at 414,217 size 50x17; Text 'Störung'
      Visibility <- "Störung_15"
   Ellipse "Ellipse_11" at 377,177 size 9x9
      Visibility <- "Störung_15"
   Ellipse "Ellipse_12" at 376,222 size 9x9
      Visibility <- "Störung_15"
   TextField "Textfeld_56" at 518,271 size 50x17; Text 'Störung'
      Visibility <- "Störung_5"
   Ellipse "Ellipse_13" at 502,276 size 9x9
      Visibility <- "Störung_5"
   Ellipse "Ellipse_14" at 376,271 size 9x9
      Visibility <- "Störung_10"
   TextField "Textfeld_57" at 322,244 size 50x17; Text 'Störung'
      Visibility <- "Störung_12"
   TextField "Textfeld_58" at 322,244 size 50x17; Text 'Störung'
      Visibility <- "Störung_13"
   Ellipse "Ellipse_15" at 336,228 size 9x9
      Visibility <- "Störung_13"
   Ellipse "Ellipse_16" at 357,228 size 9x9
      Visibility <- "Störung_12"
   TextField "Textfeld_59" at 261,244 size 50x17; Text 'Störung'
      Visibility <- "Störung_14"
   Ellipse "Ellipse_17" at 298,213 size 9x9
      Visibility <- "Störung_15"
   Ellipse "Ellipse_18" at 299,228 size 9x9
      Visibility <- "Störung_14"
   TextField "Textfeld_60" at 260,186 size 50x17; Text 'Störung'
      Visibility <- "Störung_15"
   Button "Schaltfläche_2" at 598,296 size 182x69; TextOff 'STOP ALL'
      Appearance <- "Haupt_Stop_HMI"
      on Press: SetBit("Haupt_Stop_HMI")
      on Release: ResetBit("Haupt_Stop_HMI")
   TextField "Textfeld_1" at 295,86 size 206x23; Text 'ANLAGE LÄUFT NORMAL'
      Visibility <- "GDB_PLC_Start_Modus"
   TextField "Textfeld_2" at 276,110 size 137x20; Text 'Produktion läuft seit'
      Visibility <- "GDB_PLC_Start_Modus"
   TextField "Textfeld_3" at 439,110 size 23x20; Text 'St.'
      Visibility <- "GDB_PLC_Start_Modus"
   TextField "Textfeld_7" at 488,110 size 31x20; Text 'Min.'
      Visibility <- "GDB_PLC_Start_Modus"
   IOField "EA-Feld_10" at 415,106 size 26x29; FormatPattern 99
      ProcessValue <- "GDB_PLC_Run_Hours"
      Visibility <- "GDB_PLC_Start_Modus"
   IOField "EA-Feld_11" at 462,104 size 26x32; FormatPattern 99
      ProcessValue <- "GDB_PLC_Run_Minutes"
      Visibility <- "GDB_PLC_Start_Modus"
   TextField "Textfeld_8" at 540,110 size 32x20; Text 'Sec.'
      Visibility <- "GDB_PLC_Start_Modus"
   IOField "EA-Feld_12" at 514,104 size 26x32; FormatPattern 99
      ProcessValue <- "GDB_PLC_Run_Seconds"
      Visibility <- "GDB_PLC_Start_Modus"
   Rectangle "Rechteck_8" at 8,76 size 786x61
      Visibility <- "GDB_PLC_Not_Aus_Modus"
   TextField "Textfeld_34" at 352,94 size 79x23; Text 'NOT AUS'
      Visibility <- "GDB_PLC_Not_Aus_Modus"
   Rectangle "Rechteck_9" at 7,76 size 786x61
      Visibility <- "GDB_PLC_Stop_Modus"
   TextField "Textfeld_35" at 294,95 size 165x23; Text 'ANLAGE GESTOPPT'
      Visibility <- "GDB_PLC_Stop_Modus"
   Ellipse "Ellipse_3" at 432,380 size 9x9
      Visibility <- "Störung_1"
   TextField "Textfeld_38" at 380,375 size 50x17; Text 'Störung'
      Visibility <- "Störung_1"
   Ellipse "Ellipse_5" at 509,338 size 9x9
      Visibility <- "Störung_2"
   TextField "Textfeld_40" at 522,333 size 50x17; Text 'Störung'
      Visibility <- "Störung_2"
   Ellipse "Ellipse_1" at 433,338 size 9x9
      Visibility <- "Störung_0"
   TextField "Textfeld_36" at 381,333 size 50x17; Text 'Störung'
      Visibility <- "Störung_0"
   Ellipse "Ellipse_2" at 432,300 size 9x9
      Visibility <- "Störung_3"
   TextField "Textfeld_37" at 380,295 size 50x17; Text 'Störung'
      Visibility <- "Störung_3"
   Ellipse "Ellipse_4" at 505,294 size 9x9
      Visibility <- "Störung_4"
   TextField "Textfeld_39" at 518,289 size 50x17; Text 'Störung'
      Visibility <- "Störung_4"
   TextField "Textfeld_54" at 413,255 size 50x17; Text 'Störung'
      Visibility <- "Störung_8"
   Ellipse "Ellipse_8" at 434,274 size 9x9
      Visibility <- "Störung_8"

scheduled task "Get_User"
   on Action: function_f41c6f6c("Benutzername")
*)